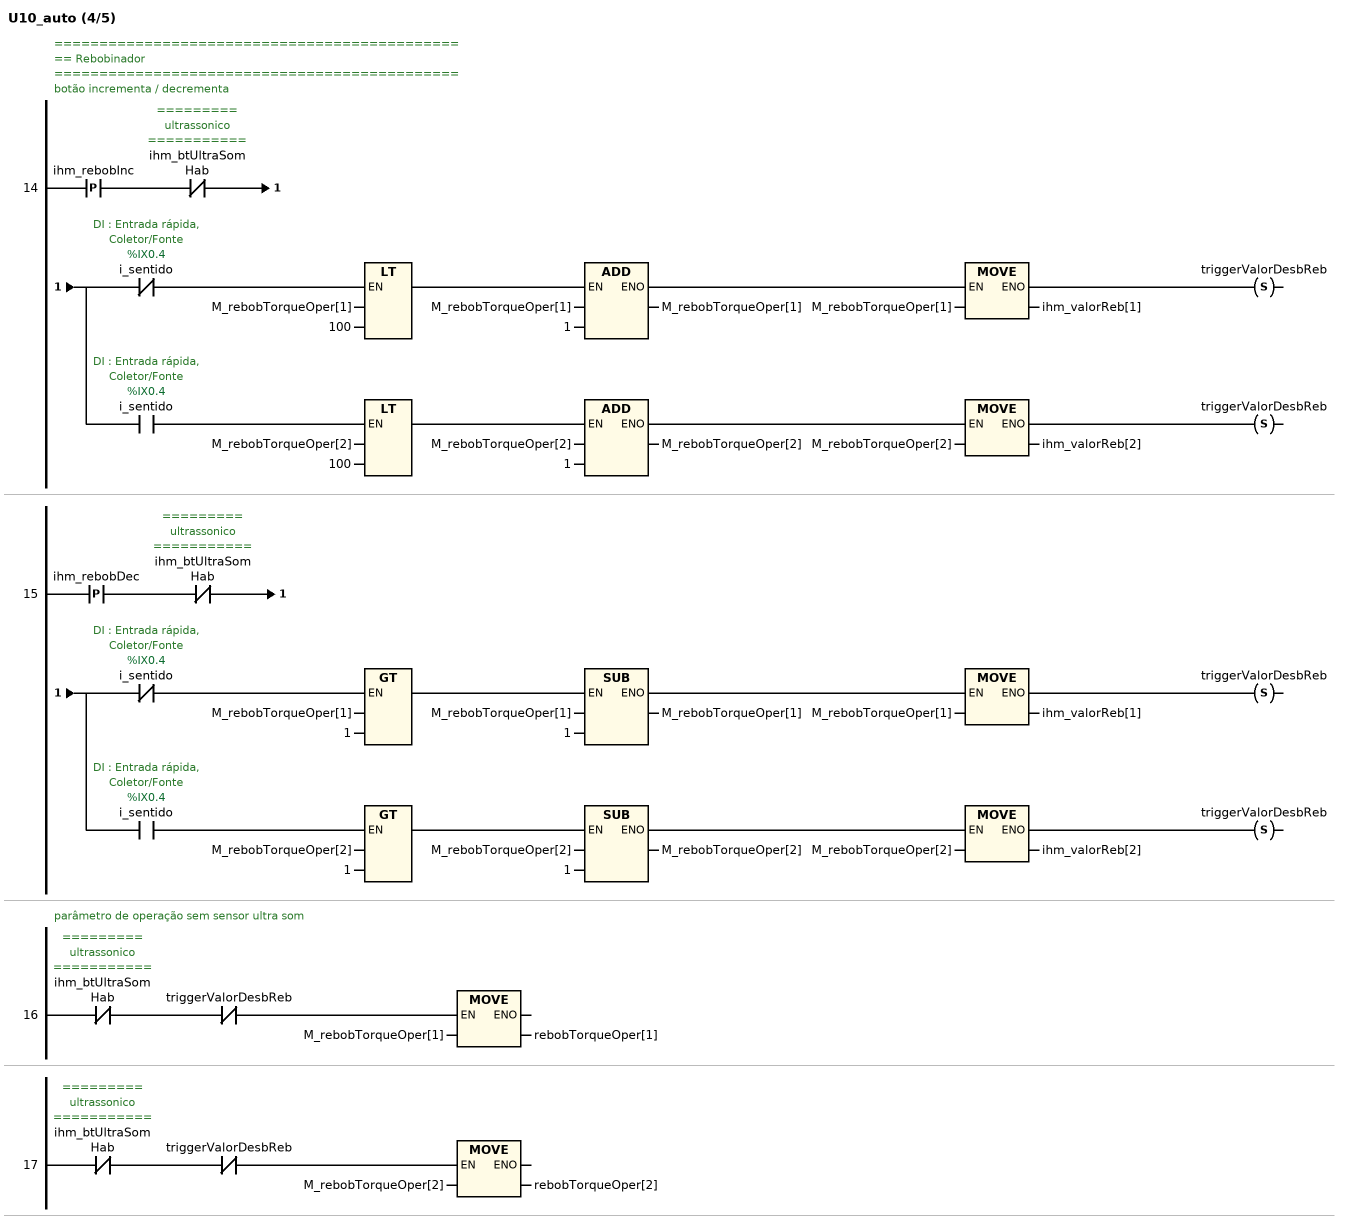
// NETWORK 14
// =============================================
// == Rebobinador
// =============================================
// botão incrementa / decrementa
//   ihm_btUltraSomHab: ========= ultrassonico ===========
//   i_sentido: DI : Entrada rápida, Coletor/Fonte | AT %IX0.4
_rt3(CLK := ihm_rebobInc);
_w7 := _rt3.Q AND NOT ihm_btUltraSomHab;
IF _w7 AND NOT i_sentido AND M_rebobTorqueOper[1] < 100 THEN
    M_rebobTorqueOper[1] := M_rebobTorqueOper[1] + 1;
END_IF
IF _w7 AND NOT i_sentido AND M_rebobTorqueOper[1] < 100 THEN ihm_valorReb[1] := M_rebobTorqueOper[1]; END_IF
triggerValorDesbReb S= _w7 AND NOT i_sentido AND M_rebobTorqueOper[1] < 100;
IF _w7 AND i_sentido AND M_rebobTorqueOper[2] < 100 THEN M_rebobTorqueOper[2] := M_rebobTorqueOper[2] + 1; END_IF
IF _w7 AND i_sentido AND M_rebobTorqueOper[2] < 100 THEN ihm_valorReb[2] := M_rebobTorqueOper[2]; END_IF
triggerValorDesbReb S= _w7 AND i_sentido AND M_rebobTorqueOper[2] < 100;

// NETWORK 15
//   ihm_btUltraSomHab: ========= ultrassonico ===========
//   i_sentido: DI : Entrada rápida, Coletor/Fonte | AT %IX0.4
_rt4(CLK := ihm_rebobDec);
_w8 := _rt4.Q AND NOT ihm_btUltraSomHab;
IF _w8 AND NOT i_sentido AND M_rebobTorqueOper[1] > 1 THEN M_rebobTorqueOper[1] := M_rebobTorqueOper[1] - 1; END_IF
IF _w8 AND NOT i_sentido AND M_rebobTorqueOper[1] > 1 THEN ihm_valorReb[1] := M_rebobTorqueOper[1]; END_IF
triggerValorDesbReb S= _w8 AND NOT i_sentido AND M_rebobTorqueOper[1] > 1;
IF _w8 AND i_sentido AND M_rebobTorqueOper[2] > 1 THEN M_rebobTorqueOper[2] := M_rebobTorqueOper[2] - 1; END_IF
IF _w8 AND i_sentido AND M_rebobTorqueOper[2] > 1 THEN ihm_valorReb[2] := M_rebobTorqueOper[2]; END_IF
triggerValorDesbReb S= _w8 AND i_sentido AND M_rebobTorqueOper[2] > 1;

// NETWORK 16
// parâmetro de operação sem sensor ultra som
//   ihm_btUltraSomHab: ========= ultrassonico ===========
//   rebobTorqueOper[1]: =================== Ultrassonico ===================
IF NOT ihm_btUltraSomHab AND NOT triggerValorDesbReb THEN rebobTorqueOper[1] := M_rebobTorqueOper[1]; END_IF

// NETWORK 17
//   ihm_btUltraSomHab: ========= ultrassonico ===========
//   rebobTorqueOper[2]: =================== Ultrassonico ===================
IF NOT ihm_btUltraSomHab AND NOT triggerValorDesbReb THEN rebobTorqueOper[2] := M_rebobTorqueOper[2]; END_IF

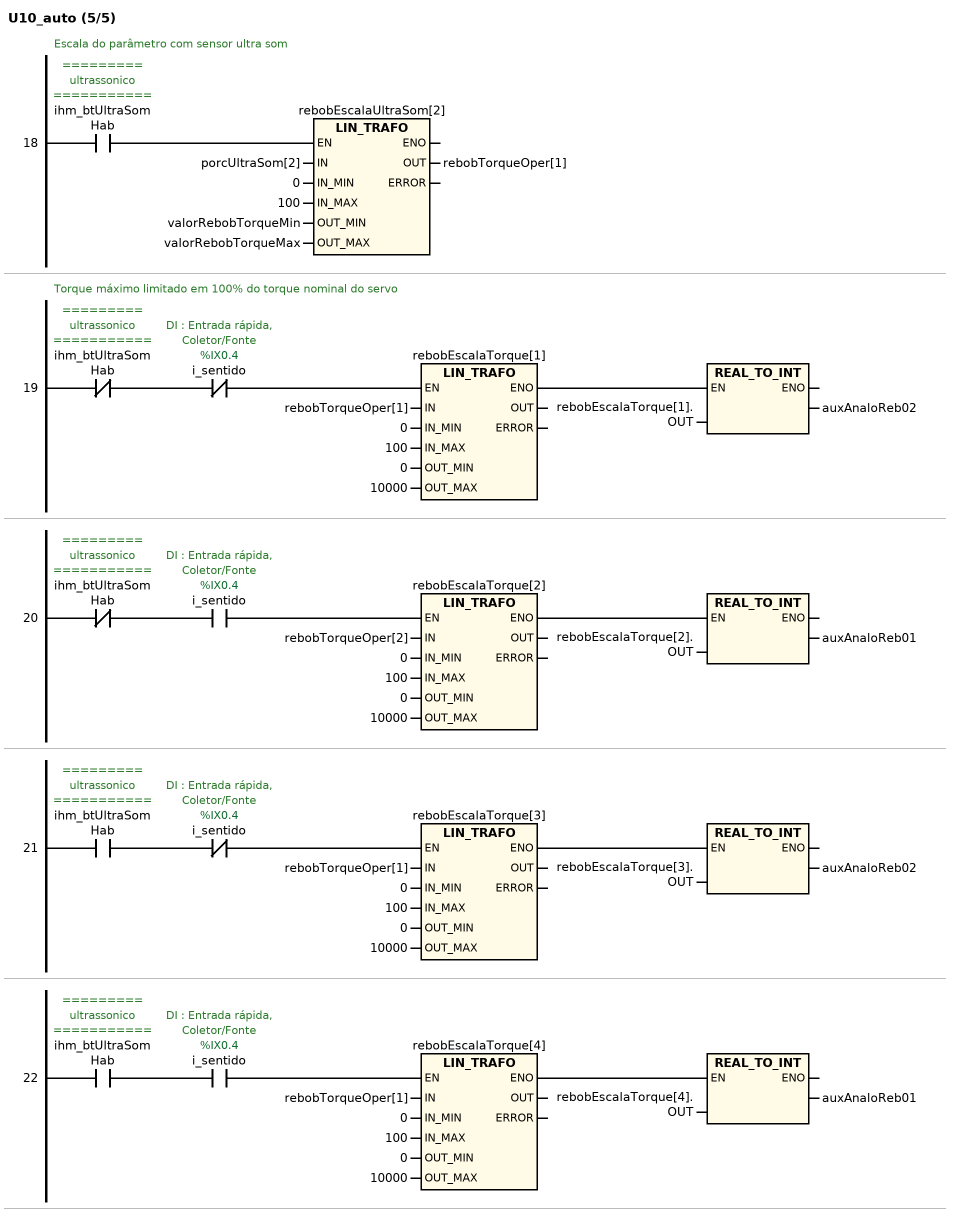
// NETWORK 18
// Escala do parâmetro com sensor ultra som
//   ihm_btUltraSomHab: ========= ultrassonico ===========
//   rebobTorqueOper[1]: =================== Ultrassonico ===================
IF ihm_btUltraSomHab THEN
    rebobEscalaUltraSom[2](
        IN := porcUltraSom[2],
        IN_MIN := 0,
        IN_MAX := 100,
        OUT_MIN := valorRebobTorqueMin,
        OUT_MAX := valorRebobTorqueMax,
        OUT => rebobTorqueOper[1]); // LIN_TRAFO
END_IF

// NETWORK 19
// Torque máximo limitado em 100% do torque nominal do servo
//   ihm_btUltraSomHab: ========= ultrassonico ===========
//   i_sentido: DI : Entrada rápida, Coletor/Fonte | AT %IX0.4
//   rebobTorqueOper[1]: =================== Ultrassonico ===================
//   rebobEscalaTorque[1].OUT: output value
_w9 := NOT ihm_btUltraSomHab AND NOT i_sentido;
IF _w9 THEN
    rebobEscalaTorque[1](IN := rebobTorqueOper[1], IN_MIN := 0, IN_MAX := 100, OUT_MIN := 0, OUT_MAX := 10000); // LIN_TRAFO
END_IF
IF _w9 THEN auxAnaloReb02 := REAL_TO_INT(rebobEscalaTorque[1].OUT); END_IF

// NETWORK 20
//   ihm_btUltraSomHab: ========= ultrassonico ===========
//   i_sentido: DI : Entrada rápida, Coletor/Fonte | AT %IX0.4
//   rebobTorqueOper[2]: =================== Ultrassonico ===================
//   rebobEscalaTorque[2].OUT: output value
_w10 := NOT ihm_btUltraSomHab AND i_sentido;
IF _w10 THEN
    rebobEscalaTorque[2](IN := rebobTorqueOper[2], IN_MIN := 0, IN_MAX := 100, OUT_MIN := 0, OUT_MAX := 10000); // LIN_TRAFO
END_IF
IF _w10 THEN auxAnaloReb01 := REAL_TO_INT(rebobEscalaTorque[2].OUT); END_IF

// NETWORK 21
//   ihm_btUltraSomHab: ========= ultrassonico ===========
//   i_sentido: DI : Entrada rápida, Coletor/Fonte | AT %IX0.4
//   rebobTorqueOper[1]: =================== Ultrassonico ===================
//   rebobEscalaTorque[3].OUT: output value
_w11 := ihm_btUltraSomHab AND NOT i_sentido;
IF _w11 THEN
    rebobEscalaTorque[3](IN := rebobTorqueOper[1], IN_MIN := 0, IN_MAX := 100, OUT_MIN := 0, OUT_MAX := 10000); // LIN_TRAFO
END_IF
IF _w11 THEN auxAnaloReb02 := REAL_TO_INT(rebobEscalaTorque[3].OUT); END_IF

// NETWORK 22
//   ihm_btUltraSomHab: ========= ultrassonico ===========
//   i_sentido: DI : Entrada rápida, Coletor/Fonte | AT %IX0.4
//   rebobTorqueOper[1]: =================== Ultrassonico ===================
//   rebobEscalaTorque[4].OUT: output value
_w12 := ihm_btUltraSomHab AND i_sentido;
IF _w12 THEN
    rebobEscalaTorque[4](IN := rebobTorqueOper[1], IN_MIN := 0, IN_MAX := 100, OUT_MIN := 0, OUT_MAX := 10000); // LIN_TRAFO
END_IF
IF _w12 THEN auxAnaloReb01 := REAL_TO_INT(rebobEscalaTorque[4].OUT); END_IF

END_PROGRAM

// MyController/Application/05_IHM/I01_geral
PROGRAM I01_geral
VAR
	auxBit				: BOOL;
END_VAR
VAR // added by the converter: edge detectors and wires of the graphical bodies
    _rt1 : R_TRIG;
END_VAR

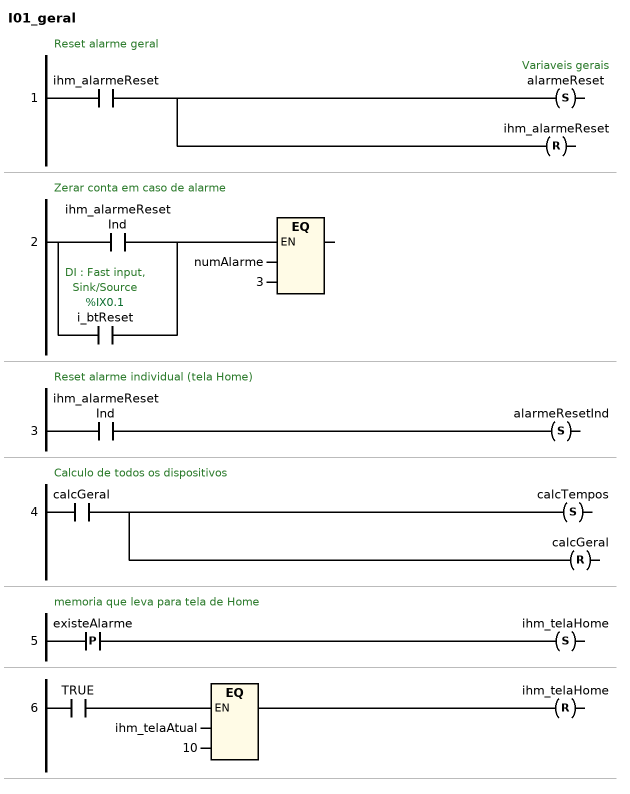
// NETWORK 1
// Reset alarme geral
//   alarmeReset: Variaveis gerais
alarmeReset S= ihm_alarmeReset;
ihm_alarmeReset R= ihm_alarmeReset;

// NETWORK 2
// Zerar conta em caso de alarme
//   i_btReset: DI : Fast input, Sink/Source | AT %IX0.1
(* (ihm_alarmeResetInd OR i_btReset) AND numAlarme = 3; result not used *)

// NETWORK 3
// Reset alarme individual (tela Home)
alarmeResetInd S= ihm_alarmeResetInd;

// NETWORK 4
// Calculo de todos os dispositivos
calcTempos S= calcGeral;
calcGeral R= calcGeral;

// NETWORK 5
// memoria que leva para tela de Home
_rt1(CLK := existeAlarme);
ihm_telaHome S= _rt1.Q;

// NETWORK 6
ihm_telaHome R= ihm_telaAtual = 10;

END_PROGRAM

// MyController/Application/05_IHM/I02_alarmes
PROGRAM I02_alarmes
VAR
	auxExisteAlarme					: BOOL;
	delayAlarme						: TON;
	memAlarme						: ARRAY[0..99] OF BOOL;
	p0								: SINT;
END_VAR


CASE alarmes.Fase OF
(*====================================
  ==  Fase 0 - alarmes 1 a 50 (0 não existe)
  ====================================*)
0:
	auxExisteAlarme:= FALSE;
	FOR p0:= 1 TO 50 DO
		IF alarme[p0] THEN
			memAlarme[p0]:= TRUE;
			auxExisteAlarme:= TRUE;
			
			IF numAlarme = 0 THEN
				numAlarme:= p0;				// pega o numero do primeiro alarme que ocorre
			END_IF
		END_IF
		
		IF numAlarme = p0 THEN
			IF alarme[p0] = 0 THEN			// verifica se o alarme que ocorreu continua ativo
				numAlarme:= 0;
			END_IF
		END_IF
	END_FOR
	alarmes.Fase:= 10;

	
(*====================================
  ==  Fase 10 - passa alarmes para ihm	
  ====================================*)
10:
	FOR p0:= 1 TO 50 DO
		ihm_alarme[p0]:= memAlarme[p0];
		memAlarme[p0]:= FALSE;
	END_FOR
	alarmes.Fase:= 11;
	
	
(*====================================
  ==  Fase 11 - verifica cancela alarmes pela IHM
  ====================================*)	
11:
	existeAlarme:= auxExisteAlarme;
	IF alarmeReset THEN
		alarmes.Fase:= 12;
	ELSE
		IF alarmeResetInd OR (i_btReset AND comando.DN) THEN
			alarme[numAlarme]:= FALSE;
			alarmeResetInd:= FALSE;
		END_IF
		alarmes.Fase:= 0;
	END_IF

	
(*====================================
  ==  Fase 12 - cancela alarmes	
  ====================================*)
12:
	alarmeReset:= FALSE;
	FOR p0:= 1 TO 50 DO
		alarme[p0]:= 0;
	END_FOR
	alarmes.Fase:= 13;
	

(*====================================
  ==  Fase 13 - espera 100ms para atualização dos bits de alarmes pelo controle
  ====================================*)	
13:
	IF delayAlarme.Q THEN
		alarmes.Fase:= 0;
	END_IF
	delayAlarme(IN:= alarmes.Fase= 13, PT:= T#100MS);

END_CASE

END_PROGRAM

// MyController/Application/05_IHM/I03_mensagens
PROGRAM I03_mensagens
VAR
	delayMensag						: TON;
	mensagens						: _exec_bits;
	p1								: DINT;
END_VAR


IF NOT mensagens.RQ THEN
	FOR p1:= 1 TO 50 DO
		IF mensagem[p1] = TRUE THEN
			mensagem[p1]:= 0;
			ihm_mensagem:= p1;
			mensagens.RQ:= TRUE;
		END_IF
	END_FOR
END_IF


// Tempo de cada mensagem na tela
delayMensag(IN := ihm_bannerMensagem, PT:= T#2500MS);
IF delayMensag.Q THEN
	mensagens.RQ:= FALSE;
	ihm_mensagem:= 0;
END_IF


ihm_bannerMensagem:= mensagens.RQ AND NOT ihm_bannerConfirma;

END_PROGRAM

// MyController/Application/05_IHM/I06_textoConfirma
PROGRAM I06_textoConfirma
VAR
END_VAR
VAR // added by the converter: edge detectors and wires of the graphical bodies
    _w1 : BOOL;
END_VAR

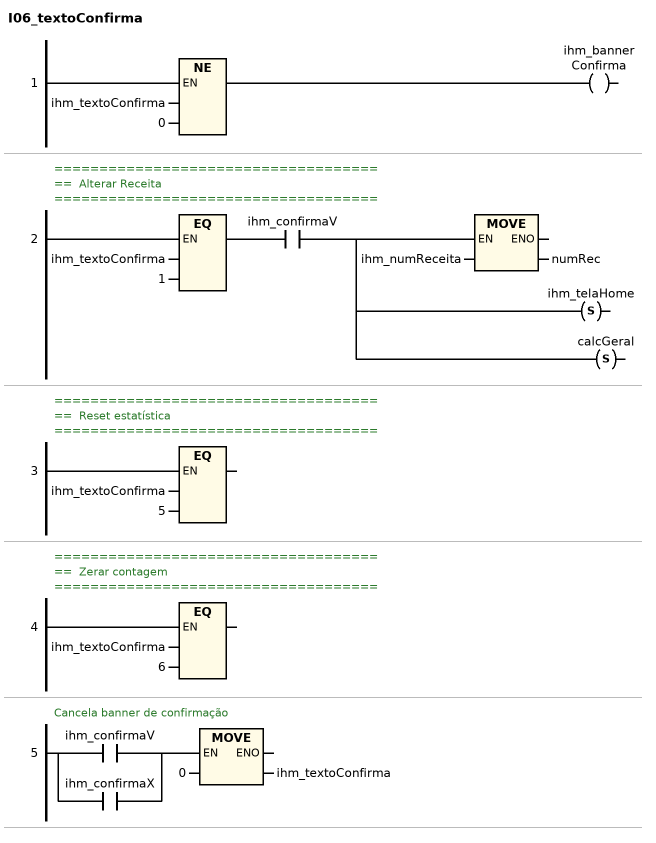
// NETWORK 1
ihm_bannerConfirma := ihm_textoConfirma <> 0;

// NETWORK 2
// ====================================
// ==  Alterar Receita
// ====================================
_w1 := ihm_textoConfirma = 1 AND ihm_confirmaV;
IF _w1 THEN numRec := ihm_numReceita; END_IF
ihm_telaHome S= _w1;
calcGeral S= _w1;

// NETWORK 3
// ====================================
// ==  Reset estatística
// ====================================
(* ihm_textoConfirma = 5; result not used *)

// NETWORK 4
// ====================================
// ==  Zerar contagem
// ====================================
(* ihm_textoConfirma = 6; result not used *)

// NETWORK 5
// Cancela banner de confirmação
IF ihm_confirmaV OR ihm_confirmaX THEN ihm_textoConfirma := 0; END_IF

END_PROGRAM

// MyController/Application/10_Relogio/AjustaDataHora
PROGRAM AjustaDataHora
VAR
	writeDateTime			: SetDateAndTime;
	readDateTime			: GetDateAndTime;
	bitScan					: BOOL;
	comOk					: BOOL;
	T_com					: TON;
END_VAR
VAR // added by the converter: edge detectors and wires of the graphical bodies
    _rt1 : R_TRIG;
END_VAR

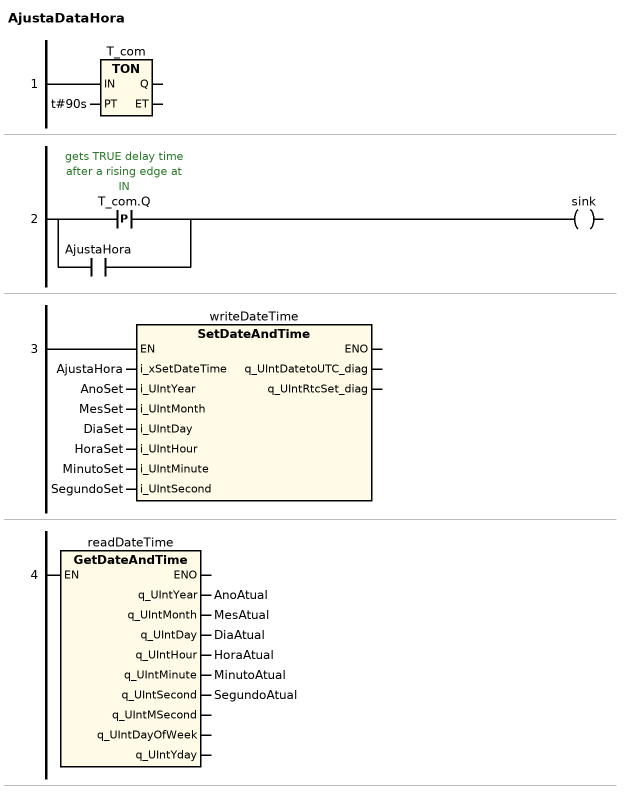
// NETWORK 1
T_com(IN := TRUE, PT := t#90s); // TON

// NETWORK 2
//   T_com.Q: gets TRUE delay time after a rising edge at IN
_rt1(CLK := T_com.Q);
sink := _rt1.Q OR AjustaHora;

// NETWORK 3
//   AnoSet: Sincroniza e ajusta o relógio da IHM
writeDateTime(
    i_xSetDateTime := AjustaHora,
    i_UIntYear := AnoSet,
    i_UIntMonth := MesSet,
    i_UIntDay := DiaSet,
    i_UIntHour := HoraSet,
    i_UIntMinute := MinutoSet,
    i_UIntSecond := SegundoSet); // SetDateAndTime

// NETWORK 4
readDateTime(
    q_UIntYear => AnoAtual,
    q_UIntMonth => MesAtual,
    q_UIntDay => DiaAtual,
    q_UIntHour => HoraAtual,
    q_UIntMinute => MinutoAtual,
    q_UIntSecond => SegundoAtual); // GetDateAndTime

END_PROGRAM

// MyController/Application/10_Relogio/SetDateAndTime
FUNCTION_BLOCK SetDateAndTime
VAR_INPUT
	i_xSetDateTime			: BOOL; (* seta novo horário na transição false para true*)
	i_UIntYear				: UINT:=2011; (*Valor para o ano a ser ajustado*)
	i_UIntMonth				: UINT:=1;(*Valor para o mes a ser ajustado*) 
	i_UIntDay				: UINT:=1;(*Valor para o dia a ser ajustado*) 
	i_UIntHour				: UINT:=0; (*Valor para a hora a ser ajustada*)
	i_UIntMinute			: UINT:=0; (*Valor para o minuto a ser ajustado*)
	i_UIntSecond			: UINT:=0;(*Valor para o segundo a ser ajustado*)
END_VAR
VAR_OUTPUT
	q_UIntDatetoUTC_diag	: UDINT; (*Status quando se =0 ok se <>0 erro nas informações de entrada*)
	q_UIntRtcSet_diag		: UDINT; (*Status quando se =0 ok se <>0 erro nas informações de entrada*)
END_VAR
VAR
	My_UTC					: DWORD; 
	MyDateTime				: SYSTIMEDATE; 
	milesec					: UINT:=0;
	dayOfWeek				: UINT:=1;
	yday					: UINT:=1;
END_VAR
VAR // added by the converter: edge detectors and wires of the graphical bodies
    _s1 : SYSTIMEDATE;
    _w1, _w2 : ANY;
END_VAR

// compose _s1 : SYSTIMEDATE
_s1.wYear := i_UIntYear;
_s1.wMonth := i_UIntMonth;
_s1.wDay := i_UIntDay;
_s1.wHour := i_UIntHour;
_s1.wMinute := i_UIntMinute;
_s1.wSecond := i_UIntSecond;
_s1.wMilliseconds := milesec;
_s1.wDayOfWeek := dayOfWeek;
_s1.wYday := yday;
MyDateTime := _s1;
_w1 := SysTimeRtcConvertDateToUtc(pDate := MyDateTime, pdwTimestampUtc := My_UTC);
q_UIntDatetoUTC_diag := _w1;
IF My_UTC <> 16#FFFFFFFF AND i_xSetDateTime THEN _w2 := SysTimeRtcSet(ulTimestamp := My_UTC); END_IF
q_UIntRtcSet_diag := _w2;
i_xSetDateTime := FALSE;

END_FUNCTION_BLOCK

// MyController/Application/10_Relogio/GetDateAndTime
FUNCTION_BLOCK GetDateAndTime
VAR_INPUT
END_VAR
VAR_OUTPUT
	q_UIntYear			: UINT; 
	q_UIntMonth			: UINT; 
	q_UIntDay			: UINT; 
	q_UIntHour			: UINT; 
	q_UIntMinute		: UINT; 
	q_UIntSecond		: UINT; 
	q_UIntMSecond		: UINT; 
	q_UIntDayOfWeek		: UINT; 
	q_UIntYday			: UINT;
END_VAR
VAR
	Ctrl_DateTime		: SYSTIMEDATE; 
	// SysTimeRtcGet operation diag 
	GetTimeResult		: UDINT; 
// SysTimeRtcConvertUtcToDate operation diag 
	UTCtoDate_diag		: UDINT; 
END_VAR
VAR // added by the converter: edge detectors and wires of the graphical bodies
    _w1, _w2 : ANY;
END_VAR

_w1 := SysTimeRtcGet(pResult := GetTimeResult);
_w2 := SysTimeRtcConvertUtcToDate(dwTimestampUtc := _w1, pDate := Ctrl_DateTime);
UTCtoDate_diag := _w2;
q_UIntYear := Ctrl_DateTime.SYSTIMEDATE;
q_UIntMonth := Ctrl_DateTime.wYear;
q_UIntDay := Ctrl_DateTime.wMonth;
q_UIntHour := Ctrl_DateTime.wDay;
q_UIntMinute := Ctrl_DateTime.wHour;
q_UIntSecond := Ctrl_DateTime.wMinute;
q_UIntMSecond := Ctrl_DateTime.wSecond;
q_UIntDayOfWeek := Ctrl_DateTime.wMilliseconds;
q_UIntYday := Ctrl_DateTime.wDayOfWeek;

END_FUNCTION_BLOCK

// MyController/Application/02_Rebobinadores/RB01_enableReb
PROGRAM RB01_enableReb
VAR
	TL_Rebobinadores 			 	: TON;
	TL_delayTorque					: ARRAY [0..1] OF TON;
	auxDesligaReb					: BOOL;
END_VAR
VAR // added by the converter: edge detectors and wires of the graphical bodies
    _rt1 : R_TRIG;
    _ft1 : F_TRIG;
    _w1 : BOOL;
END_VAR

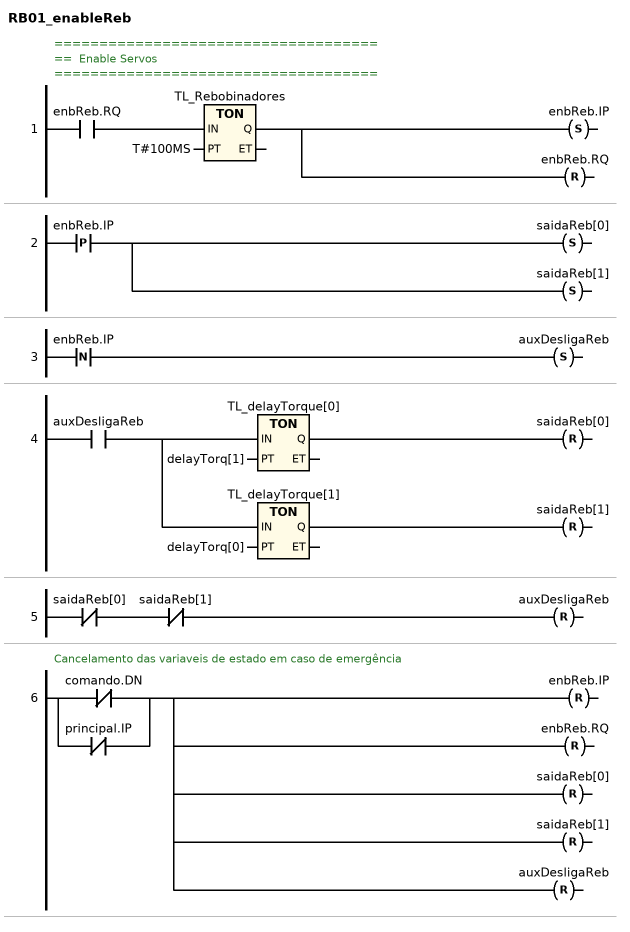
// NETWORK 1
// ====================================
// ==  Enable Servos
// ====================================
TL_Rebobinadores(IN := enbReb.RQ, PT := T#100MS); // TON
enbReb.IP S= TL_Rebobinadores.Q;
enbReb.RQ R= TL_Rebobinadores.Q;

// NETWORK 2
_rt1(CLK := enbReb.IP);
saidaReb[0] S= _rt1.Q;
saidaReb[1] S= _rt1.Q;

// NETWORK 3
_ft1(CLK := enbReb.IP);
auxDesligaReb S= _ft1.Q;

// NETWORK 4
TL_delayTorque[0](IN := auxDesligaReb, PT := delayTorq[1]); // TON
saidaReb[0] R= TL_delayTorque[0].Q;
TL_delayTorque[1](IN := auxDesligaReb, PT := delayTorq[0]); // TON
saidaReb[1] R= TL_delayTorque[1].Q;

// NETWORK 5
auxDesligaReb R= NOT saidaReb[0] AND NOT saidaReb[1];

// NETWORK 6
// Cancelamento das variaveis de estado em caso de emergência
_w1 := NOT comando.DN OR NOT principal.IP;
enbReb.IP R= _w1;
enbReb.RQ R= _w1;
saidaReb[0] R= _w1;
saidaReb[1] R= _w1;
auxDesligaReb R= _w1;

END_PROGRAM

// MyController/Application/11_FB/RTO
FUNCTION_BLOCK RTO
VAR_INPUT
	IN				: BOOL;
	PT				: TIME;
	RST				: BOOL;
END_VAR
VAR_OUTPUT
	Q				: BOOL;
	ACC				: TIME;
END_VAR
VAR
	auxIn			: BOOL;
	auxAcc			: TIME;
	timer			: TON;
END_VAR

IF IN AND NOT Q THEN
    ACC:= auxAcc + timer.ET;
    auxIn:= true;
end_if;

if not IN then
    auxAcc:= ACC;
    auxIn:= false;
end_if;

if ACC >= PT then
    Q:= true;
    ACC:= PT;
    auxIn:= false;
end_if;

if RST then
    Q:= false;
    ACC:= T#0s;
    auxAcc:= T#0s;
    auxIn:= false;
end_if;

timer(IN:= auxIn, PT:= T#999999S);

END_FUNCTION_BLOCK
